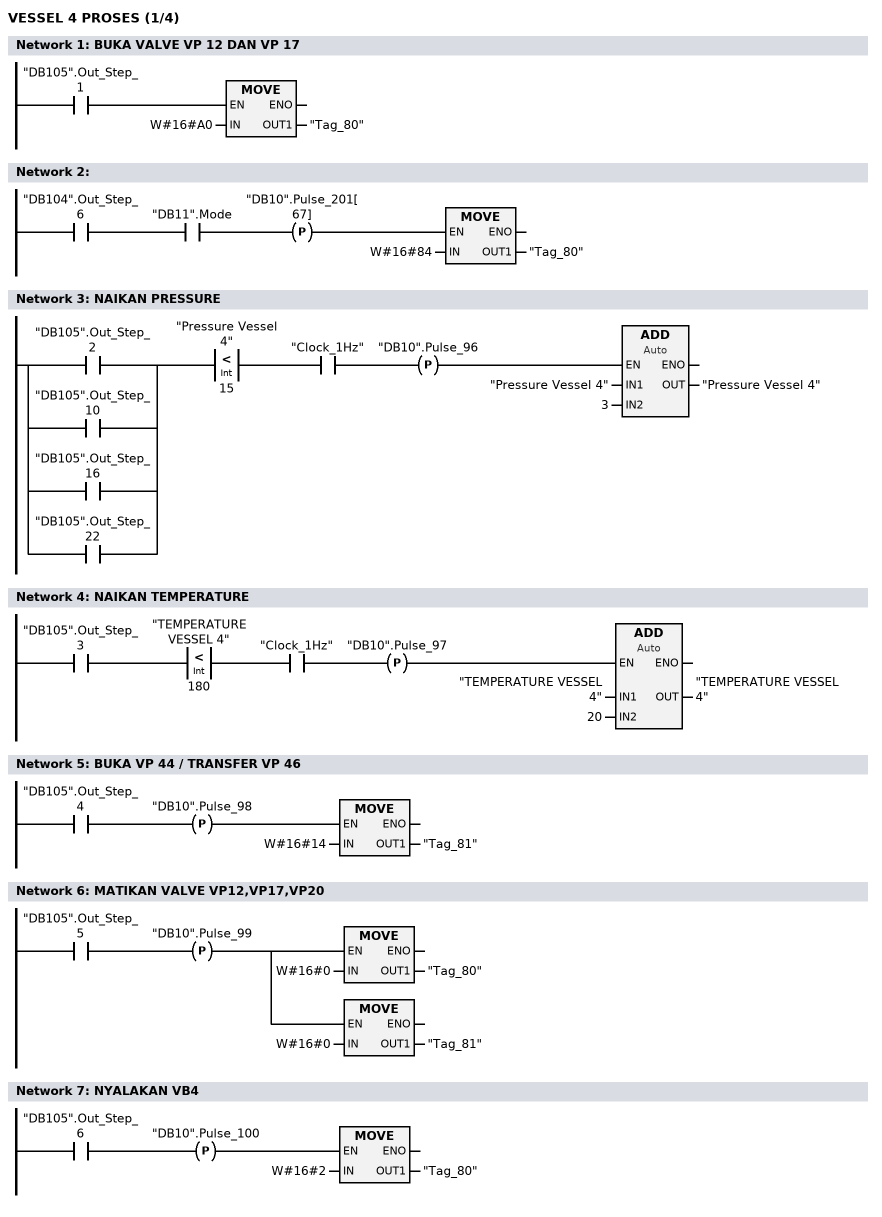
   RUNG wire#powerrail
      Contact( "DB105".Out_Step_1 )
      Move(in := W#16#A0, out1 => "Tag_80")
   END_RUNG
   // the same network as SCL:
   IF "DB105".Out_Step_1 THEN "Tag_80" := W#16#A0; END_IF;
END_REGION

REGION Network 2
   RUNG wire#powerrail
      Contact( "DB104".Out_Step_6 )
      Contact( "DB11".Mode )
      P_Trig( "DB10".Pulse_201[67] )
      Move(in := W#16#84, out1 => "Tag_80")
   END_RUNG
   // the same network as SCL:
   #_w1 := "DB104".Out_Step_6 AND "DB11".Mode;
   #_w2 := #_w1 AND NOT "DB10".Pulse_201[67];   // rising edge
   "DB10".Pulse_201[67] := #_w1;
   IF #_w2 THEN "Tag_80" := W#16#84; END_IF;
END_REGION

REGION Network 3: NAIKAN PRESSURE
   RUNG wire#powerrail
      Contact( "DB105".Out_Step_2 )
      wire#w1
      { S7_Templates := "SrcType := Int" } LT_Contact(in1 := "Pressure Vessel 4", in2 := 15)
      Contact( "Clock_1Hz" )
      P_Trig( "DB10".Pulse_96 )
      Add(in1 := "Pressure Vessel 4", in2 := 3, out => "Pressure Vessel 4")
   END_RUNG
   RUNG wire#powerrail
      Contact( "DB105".Out_Step_10 )
   END_RUNG wire#w1
   RUNG wire#powerrail
      Contact( "DB105".Out_Step_16 )
   END_RUNG wire#w1
   RUNG wire#powerrail
      Contact( "DB105".Out_Step_22 )
   END_RUNG wire#w1
   // the same network as SCL:
   #_w1 := ("DB105".Out_Step_2 OR "DB105".Out_Step_10 OR "DB105".Out_Step_16 OR "DB105".Out_Step_22) AND ("Pressure Vessel 4" < 15) AND "Clock_1Hz";
   #_w2 := #_w1 AND NOT "DB10".Pulse_96;   // rising edge
   "DB10".Pulse_96 := #_w1;
   IF #_w2 THEN "Pressure Vessel 4" := "Pressure Vessel 4" + 3; END_IF;
END_REGION

REGION Network 4: NAIKAN TEMPERATURE
   RUNG wire#powerrail
      Contact( "DB105".Out_Step_3 )
      { S7_Templates := "SrcType := Int" } LT_Contact(in1 := "TEMPERATURE VESSEL 4", in2 := 180)
      Contact( "Clock_1Hz" )
      P_Trig( "DB10".Pulse_97 )
      Add(in1 := "TEMPERATURE VESSEL 4", in2 := 20, out => "TEMPERATURE VESSEL 4")
   END_RUNG
   // the same network as SCL:
   #_w1 := "DB105".Out_Step_3 AND ("TEMPERATURE VESSEL 4" < 180) AND "Clock_1Hz";
   #_w2 := #_w1 AND NOT "DB10".Pulse_97;   // rising edge
   "DB10".Pulse_97 := #_w1;
   IF #_w2 THEN "TEMPERATURE VESSEL 4" := "TEMPERATURE VESSEL 4" + 20; END_IF;
END_REGION

REGION Network 5: BUKA VP 44 / TRANSFER VP 46
   RUNG wire#powerrail
      Contact( "DB105".Out_Step_4 )
      P_Trig( "DB10".Pulse_98 )
      Move(in := W#16#14, out1 => "Tag_81")
   END_RUNG
   // the same network as SCL:
   #_w1 := "DB105".Out_Step_4 AND NOT "DB10".Pulse_98;   // rising edge
   "DB10".Pulse_98 := "DB105".Out_Step_4;
   IF #_w1 THEN "Tag_81" := W#16#14; END_IF;
END_REGION

REGION Network 6: MATIKAN VALVE VP12,VP17,VP20
   RUNG wire#powerrail
      Contact( "DB105".Out_Step_5 )
      P_Trig( "DB10".Pulse_99 )
      wire#w1
      Move(in := W#16#0, out1 => "Tag_80")
   END_RUNG
   RUNG wire#w1
      Move(in := W#16#0, out1 => "Tag_81")
   END_RUNG
   // the same network as SCL:
   #_w1 := "DB105".Out_Step_5 AND NOT "DB10".Pulse_99;   // rising edge
   "DB10".Pulse_99 := "DB105".Out_Step_5;
   IF #_w1 THEN
       "Tag_80" := W#16#0;
       "Tag_81" := W#16#0;
   END_IF;
END_REGION

REGION Network 7: NYALAKAN VB4
   RUNG wire#powerrail
      Contact( "DB105".Out_Step_6 )
      P_Trig( "DB10".Pulse_100 )
      Move(in := W#16#2, out1 => "Tag_80")
   END_RUNG
   // the same network as SCL:
   #_w1 := "DB105".Out_Step_6 AND NOT "DB10".Pulse_100;   // rising edge
   "DB10".Pulse_100 := "DB105".Out_Step_6;
   IF #_w1 THEN "Tag_80" := W#16#2; END_IF;
END_REGION

REGION Network 8: TURUNKAN PRESSURE
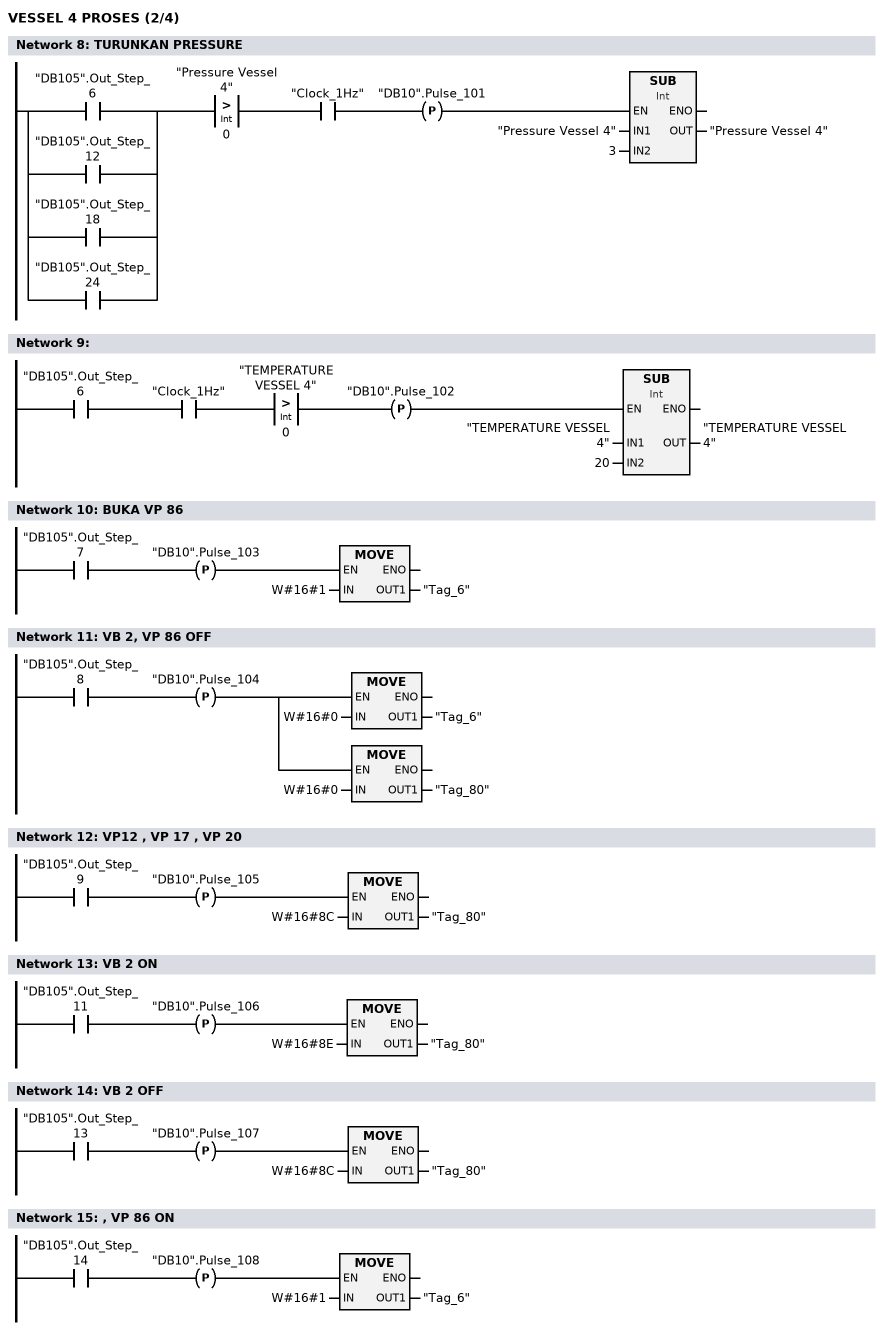
   RUNG wire#powerrail
      Contact( "DB105".Out_Step_6 )
      wire#w1
      { S7_Templates := "SrcType := Int" } GT_Contact(in1 := "Pressure Vessel 4", in2 := 0)
      Contact( "Clock_1Hz" )
      P_Trig( "DB10".Pulse_101 )
      { S7_Templates := "SrcType := Int" } Sub(in1 := "Pressure Vessel 4", in2 := 3, out => "Pressure Vessel 4")
   END_RUNG
   RUNG wire#powerrail
      Contact( "DB105".Out_Step_12 )
   END_RUNG wire#w1
   RUNG wire#powerrail
      Contact( "DB105".Out_Step_18 )
   END_RUNG wire#w1
   RUNG wire#powerrail
      Contact( "DB105".Out_Step_24 )
   END_RUNG wire#w1
   // the same network as SCL:
   #_w1 := ("DB105".Out_Step_6 OR "DB105".Out_Step_12 OR "DB105".Out_Step_18 OR "DB105".Out_Step_24) AND ("Pressure Vessel 4" > 0) AND "Clock_1Hz";
   #_w2 := #_w1 AND NOT "DB10".Pulse_101;   // rising edge
   "DB10".Pulse_101 := #_w1;
   IF #_w2 THEN "Pressure Vessel 4" := "Pressure Vessel 4" - 3; END_IF;
END_REGION

REGION Network 9
   RUNG wire#powerrail
      Contact( "DB105".Out_Step_6 )
      Contact( "Clock_1Hz" )
      { S7_Templates := "SrcType := Int" } GT_Contact(in1 := "TEMPERATURE VESSEL 4", in2 := 0)
      P_Trig( "DB10".Pulse_102 )
      { S7_Templates := "SrcType := Int" } Sub(in1 := "TEMPERATURE VESSEL 4", in2 := 20, out => "TEMPERATURE VESSEL 4")
   END_RUNG
   // the same network as SCL:
   #_w1 := "DB105".Out_Step_6 AND "Clock_1Hz" AND ("TEMPERATURE VESSEL 4" > 0);
   #_w2 := #_w1 AND NOT "DB10".Pulse_102;   // rising edge
   "DB10".Pulse_102 := #_w1;
   IF #_w2 THEN "TEMPERATURE VESSEL 4" := "TEMPERATURE VESSEL 4" - 20; END_IF;
END_REGION

REGION Network 10: BUKA VP 86
   RUNG wire#powerrail
      Contact( "DB105".Out_Step_7 )
      P_Trig( "DB10".Pulse_103 )
      Move(in := W#16#1, out1 => "Tag_6")
   END_RUNG
   // the same network as SCL:
   #_w1 := "DB105".Out_Step_7 AND NOT "DB10".Pulse_103;   // rising edge
   "DB10".Pulse_103 := "DB105".Out_Step_7;
   IF #_w1 THEN "Tag_6" := W#16#1; END_IF;
END_REGION

REGION Network 11: VB 2, VP 86 OFF
   RUNG wire#powerrail
      Contact( "DB105".Out_Step_8 )
      P_Trig( "DB10".Pulse_104 )
      wire#w1
      Move(in := W#16#0, out1 => "Tag_6")
   END_RUNG
   RUNG wire#w1
      Move(in := W#16#0, out1 => "Tag_80")
   END_RUNG
   // the same network as SCL:
   #_w1 := "DB105".Out_Step_8 AND NOT "DB10".Pulse_104;   // rising edge
   "DB10".Pulse_104 := "DB105".Out_Step_8;
   IF #_w1 THEN
       "Tag_6" := W#16#0;
       "Tag_80" := W#16#0;
   END_IF;
END_REGION

REGION Network 12: VP12 , VP 17 , VP 20
   RUNG wire#powerrail
      Contact( "DB105".Out_Step_9 )
      P_Trig( "DB10".Pulse_105 )
      Move(in := W#16#8C, out1 => "Tag_80")
   END_RUNG
   // the same network as SCL:
   #_w1 := "DB105".Out_Step_9 AND NOT "DB10".Pulse_105;   // rising edge
   "DB10".Pulse_105 := "DB105".Out_Step_9;
   IF #_w1 THEN "Tag_80" := W#16#8C; END_IF;
END_REGION

REGION Network 13: VB 2 ON
   RUNG wire#powerrail
      Contact( "DB105".Out_Step_11 )
      P_Trig( "DB10".Pulse_106 )
      Move(in := W#16#8E, out1 => "Tag_80")
   END_RUNG
   // the same network as SCL:
   #_w1 := "DB105".Out_Step_11 AND NOT "DB10".Pulse_106;   // rising edge
   "DB10".Pulse_106 := "DB105".Out_Step_11;
   IF #_w1 THEN "Tag_80" := W#16#8E; END_IF;
END_REGION

REGION Network 14: VB 2 OFF
   RUNG wire#powerrail
      Contact( "DB105".Out_Step_13 )
      P_Trig( "DB10".Pulse_107 )
      Move(in := W#16#8C, out1 => "Tag_80")
   END_RUNG
   // the same network as SCL:
   #_w1 := "DB105".Out_Step_13 AND NOT "DB10".Pulse_107;   // rising edge
   "DB10".Pulse_107 := "DB105".Out_Step_13;
   IF #_w1 THEN "Tag_80" := W#16#8C; END_IF;
END_REGION

REGION Network 15: , VP 86 ON
   RUNG wire#powerrail
      Contact( "DB105".Out_Step_14 )
      P_Trig( "DB10".Pulse_108 )
      Move(in := W#16#1, out1 => "Tag_6")
   END_RUNG
   // the same network as SCL:
   #_w1 := "DB105".Out_Step_14 AND NOT "DB10".Pulse_108;   // rising edge
   "DB10".Pulse_108 := "DB105".Out_Step_14;
   IF #_w1 THEN "Tag_6" := W#16#1; END_IF;
END_REGION

REGION Network 16: VP 86 OFF
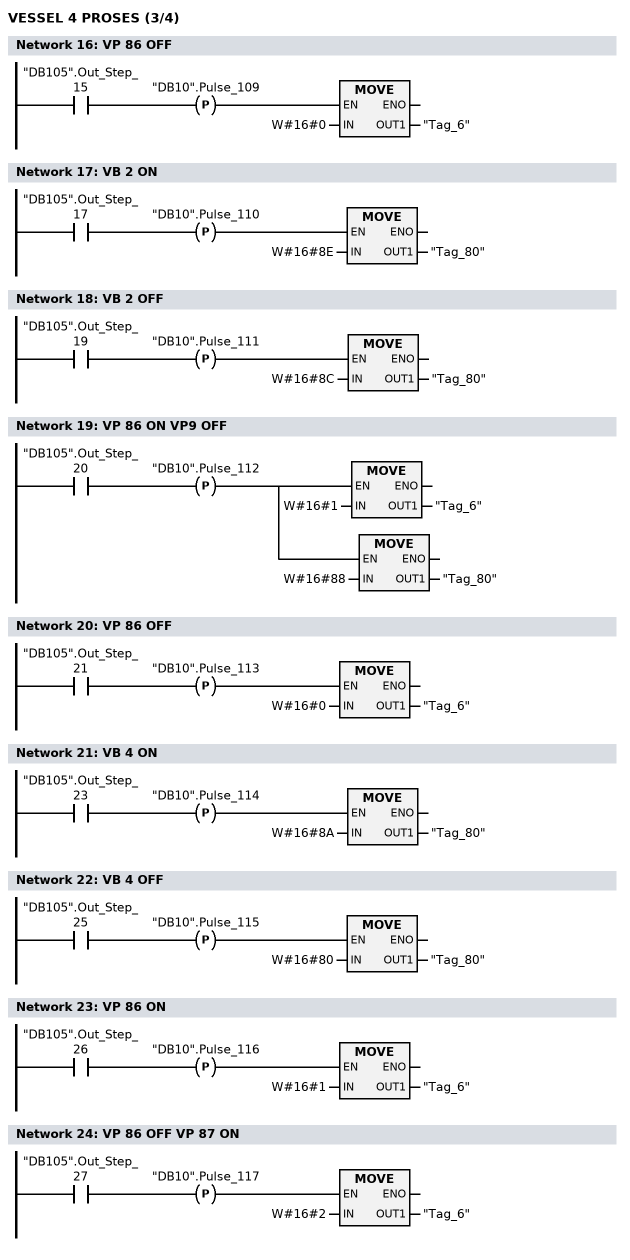
   RUNG wire#powerrail
      Contact( "DB105".Out_Step_15 )
      P_Trig( "DB10".Pulse_109 )
      Move(in := W#16#0, out1 => "Tag_6")
   END_RUNG
   // the same network as SCL:
   #_w1 := "DB105".Out_Step_15 AND NOT "DB10".Pulse_109;   // rising edge
   "DB10".Pulse_109 := "DB105".Out_Step_15;
   IF #_w1 THEN "Tag_6" := W#16#0; END_IF;
END_REGION

REGION Network 17: VB 2 ON
   RUNG wire#powerrail
      Contact( "DB105".Out_Step_17 )
      P_Trig( "DB10".Pulse_110 )
      Move(in := W#16#8E, out1 => "Tag_80")
   END_RUNG
   // the same network as SCL:
   #_w1 := "DB105".Out_Step_17 AND NOT "DB10".Pulse_110;   // rising edge
   "DB10".Pulse_110 := "DB105".Out_Step_17;
   IF #_w1 THEN "Tag_80" := W#16#8E; END_IF;
END_REGION

REGION Network 18: VB 2 OFF
   RUNG wire#powerrail
      Contact( "DB105".Out_Step_19 )
      P_Trig( "DB10".Pulse_111 )
      Move(in := W#16#8C, out1 => "Tag_80")
   END_RUNG
   // the same network as SCL:
   #_w1 := "DB105".Out_Step_19 AND NOT "DB10".Pulse_111;   // rising edge
   "DB10".Pulse_111 := "DB105".Out_Step_19;
   IF #_w1 THEN "Tag_80" := W#16#8C; END_IF;
END_REGION

REGION Network 19: VP 86 ON VP9 OFF
   RUNG wire#powerrail
      Contact( "DB105".Out_Step_20 )
      P_Trig( "DB10".Pulse_112 )
      wire#w1
      Move(in := W#16#1, out1 => "Tag_6")
   END_RUNG
   RUNG wire#w1
      Move(in := W#16#88, out1 => "Tag_80")
   END_RUNG
   // the same network as SCL:
   #_w1 := "DB105".Out_Step_20 AND NOT "DB10".Pulse_112;   // rising edge
   "DB10".Pulse_112 := "DB105".Out_Step_20;
   IF #_w1 THEN
       "Tag_6" := W#16#1;
       "Tag_80" := W#16#88;
   END_IF;
END_REGION

REGION Network 20: VP 86 OFF
   RUNG wire#powerrail
      Contact( "DB105".Out_Step_21 )
      P_Trig( "DB10".Pulse_113 )
      Move(in := W#16#0, out1 => "Tag_6")
   END_RUNG
   // the same network as SCL:
   #_w1 := "DB105".Out_Step_21 AND NOT "DB10".Pulse_113;   // rising edge
   "DB10".Pulse_113 := "DB105".Out_Step_21;
   IF #_w1 THEN "Tag_6" := W#16#0; END_IF;
END_REGION

REGION Network 21: VB 4 ON
   RUNG wire#powerrail
      Contact( "DB105".Out_Step_23 )
      P_Trig( "DB10".Pulse_114 )
      Move(in := W#16#8A, out1 => "Tag_80")
   END_RUNG
   // the same network as SCL:
   #_w1 := "DB105".Out_Step_23 AND NOT "DB10".Pulse_114;   // rising edge
   "DB10".Pulse_114 := "DB105".Out_Step_23;
   IF #_w1 THEN "Tag_80" := W#16#8A; END_IF;
END_REGION

REGION Network 22: VB 4 OFF
   RUNG wire#powerrail
      Contact( "DB105".Out_Step_25 )
      P_Trig( "DB10".Pulse_115 )
      Move(in := W#16#80, out1 => "Tag_80")
   END_RUNG
   // the same network as SCL:
   #_w1 := "DB105".Out_Step_25 AND NOT "DB10".Pulse_115;   // rising edge
   "DB10".Pulse_115 := "DB105".Out_Step_25;
   IF #_w1 THEN "Tag_80" := W#16#80; END_IF;
END_REGION

REGION Network 23: VP 86 ON
   RUNG wire#powerrail
      Contact( "DB105".Out_Step_26 )
      P_Trig( "DB10".Pulse_116 )
      Move(in := W#16#1, out1 => "Tag_6")
   END_RUNG
   // the same network as SCL:
   #_w1 := "DB105".Out_Step_26 AND NOT "DB10".Pulse_116;   // rising edge
   "DB10".Pulse_116 := "DB105".Out_Step_26;
   IF #_w1 THEN "Tag_6" := W#16#1; END_IF;
END_REGION

REGION Network 24: VP 86 OFF VP 87 ON
   RUNG wire#powerrail
      Contact( "DB105".Out_Step_27 )
      P_Trig( "DB10".Pulse_117 )
      Move(in := W#16#2, out1 => "Tag_6")
   END_RUNG
   // the same network as SCL:
   #_w1 := "DB105".Out_Step_27 AND NOT "DB10".Pulse_117;   // rising edge
   "DB10".Pulse_117 := "DB105".Out_Step_27;
   IF #_w1 THEN "Tag_6" := W#16#2; END_IF;
END_REGION

REGION Network 25: VP 87 OFF
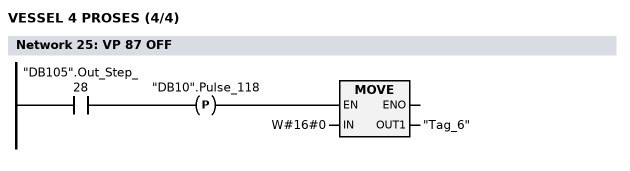
   RUNG wire#powerrail
      Contact( "DB105".Out_Step_28 )
      P_Trig( "DB10".Pulse_118 )
      Move(in := W#16#0, out1 => "Tag_6")
   END_RUNG
   // the same network as SCL:
   #_w1 := "DB105".Out_Step_28 AND NOT "DB10".Pulse_118;   // rising edge
   "DB10".Pulse_118 := "DB105".Out_Step_28;
   IF #_w1 THEN "Tag_6" := W#16#0; END_IF;
END_REGION
END_FUNCTION

FUNCTION "SEQUENCE V4 PROSES" : Void   // FC16, LAD
{ S7_Optimized_Access := 'TRUE' }
VERSION : 0.1
   VAR_TEMP   // added for the SCL form of the ladder/FBD networks
      _w1 : Bool;
      _w2 : Bool;
      _s5time1 : S5Time;
   END_VAR
BEGIN

REGION Network 1: START PROSES
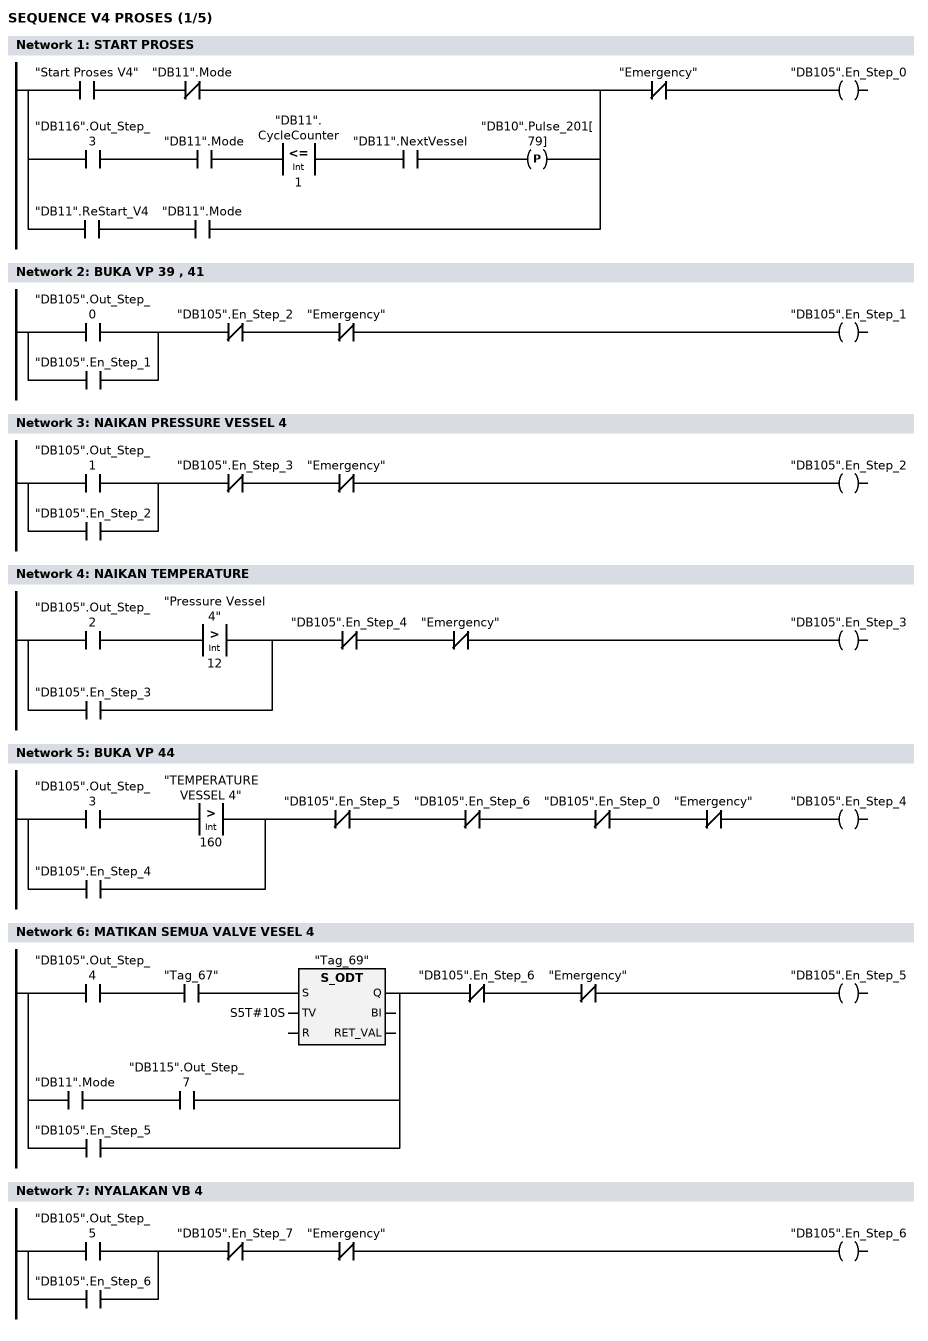
   RUNG wire#powerrail
      Contact( "Start Proses V4" )
      I_Contact( "DB11".Mode )
      wire#w1
      I_Contact( "Emergency" )
      Coil( "DB105".En_Step_0 )
   END_RUNG
   RUNG wire#powerrail
      Contact( "DB116".Out_Step_3 )
      Contact( "DB11".Mode )
      { S7_Templates := "SrcType := Int" } LE_Contact(in1 := "DB11".CycleCounter, in2 := 1)
      Contact( "DB11".NextVessel )
      P_Trig( "DB10".Pulse_201[79] )
   END_RUNG wire#w1
   RUNG wire#powerrail
      Contact( "DB11".ReStart_V4 )
      Contact( "DB11".Mode )
   END_RUNG wire#w1
   // the same network as SCL:
   #_w1 := "DB116".Out_Step_3 AND "DB11".Mode AND ("DB11".CycleCounter <= 1) AND "DB11".NextVessel;
   #_w2 := #_w1 AND NOT "DB10".Pulse_201[79];   // rising edge
   "DB10".Pulse_201[79] := #_w1;
   "DB105".En_Step_0 := (("Start Proses V4" AND NOT "DB11".Mode) OR #_w2 OR ("DB11".ReStart_V4 AND "DB11".Mode)) AND NOT "Emergency";
END_REGION

REGION Network 2: BUKA VP 39 , 41
   RUNG wire#powerrail
      Contact( "DB105".Out_Step_0 )
      wire#w1
      I_Contact( "DB105".En_Step_2 )
      I_Contact( "Emergency" )
      Coil( "DB105".En_Step_1 )
   END_RUNG
   RUNG wire#powerrail
      Contact( "DB105".En_Step_1 )
   END_RUNG wire#w1
   // the same network as SCL:
   "DB105".En_Step_1 := ("DB105".Out_Step_0 OR "DB105".En_Step_1) AND NOT "DB105".En_Step_2 AND NOT "Emergency";
END_REGION

REGION Network 3: NAIKAN PRESSURE VESSEL 4
   RUNG wire#powerrail
      Contact( "DB105".Out_Step_1 )
      wire#w1
      I_Contact( "DB105".En_Step_3 )
      I_Contact( "Emergency" )
      Coil( "DB105".En_Step_2 )
   END_RUNG
   RUNG wire#powerrail
      Contact( "DB105".En_Step_2 )
   END_RUNG wire#w1
   // the same network as SCL:
   "DB105".En_Step_2 := ("DB105".Out_Step_1 OR "DB105".En_Step_2) AND NOT "DB105".En_Step_3 AND NOT "Emergency";
END_REGION

REGION Network 4: NAIKAN TEMPERATURE
   RUNG wire#powerrail
      Contact( "DB105".Out_Step_2 )
      { S7_Templates := "SrcType := Int" } GT_Contact(in1 := "Pressure Vessel 4", in2 := 12)
      wire#w1
      I_Contact( "DB105".En_Step_4 )
      I_Contact( "Emergency" )
      Coil( "DB105".En_Step_3 )
   END_RUNG
   RUNG wire#powerrail
      Contact( "DB105".En_Step_3 )
   END_RUNG wire#w1
   // the same network as SCL:
   "DB105".En_Step_3 := (("DB105".Out_Step_2 AND ("Pressure Vessel 4" > 12)) OR "DB105".En_Step_3) AND NOT "DB105".En_Step_4 AND NOT "Emergency";
END_REGION

REGION Network 5: BUKA VP 44
   RUNG wire#powerrail
      Contact( "DB105".Out_Step_3 )
      { S7_Templates := "SrcType := Int" } GT_Contact(in1 := "TEMPERATURE VESSEL 4", in2 := 160)
      wire#w1
      I_Contact( "DB105".En_Step_5 )
      I_Contact( "DB105".En_Step_6 )
      I_Contact( "DB105".En_Step_0 )
      I_Contact( "Emergency" )
      Coil( "DB105".En_Step_4 )
   END_RUNG
   RUNG wire#powerrail
      Contact( "DB105".En_Step_4 )
   END_RUNG wire#w1
   // the same network as SCL:
   "DB105".En_Step_4 := (("DB105".Out_Step_3 AND ("TEMPERATURE VESSEL 4" > 160)) OR "DB105".En_Step_4) AND NOT "DB105".En_Step_5 AND NOT "DB105".En_Step_6 AND NOT "DB105".En_Step_0 AND NOT "Emergency";
END_REGION

REGION Network 6: MATIKAN SEMUA VALVE VESEL 4
   RUNG wire#powerrail
      Contact( "DB105".Out_Step_4 )
      Contact( "Tag_67" )
      S_ODT(T_NO := "Tag_69", TV := S5T#10S, R :=, BI =>, RET_VAL =>)
      wire#w1
      I_Contact( "DB105".En_Step_6 )
      I_Contact( "Emergency" )
      Coil( "DB105".En_Step_5 )
   END_RUNG
   RUNG wire#powerrail
      Contact( "DB11".Mode )
      Contact( "DB115".Out_Step_7 )
   END_RUNG wire#w1
   RUNG wire#powerrail
      Contact( "DB105".En_Step_5 )
   END_RUNG wire#w1
   // the same network as SCL:
   #_s5time1 := S_ODT(T_NO := "Tag_69", S := "DB105".Out_Step_4 AND "Tag_67", TV := S5T#10S, Q => #_w1);
   "DB105".En_Step_5 := (#_w1 OR ("DB11".Mode AND "DB115".Out_Step_7) OR "DB105".En_Step_5) AND NOT "DB105".En_Step_6 AND NOT "Emergency";
END_REGION

REGION Network 7: NYALAKAN VB 4
   RUNG wire#powerrail
      Contact( "DB105".Out_Step_5 )
      wire#w1
      I_Contact( "DB105".En_Step_7 )
      I_Contact( "Emergency" )
      Coil( "DB105".En_Step_6 )
   END_RUNG
   RUNG wire#powerrail
      Contact( "DB105".En_Step_6 )
   END_RUNG wire#w1
   // the same network as SCL:
   "DB105".En_Step_6 := ("DB105".Out_Step_5 OR "DB105".En_Step_6) AND NOT "DB105".En_Step_7 AND NOT "Emergency";
END_REGION

REGION Network 8
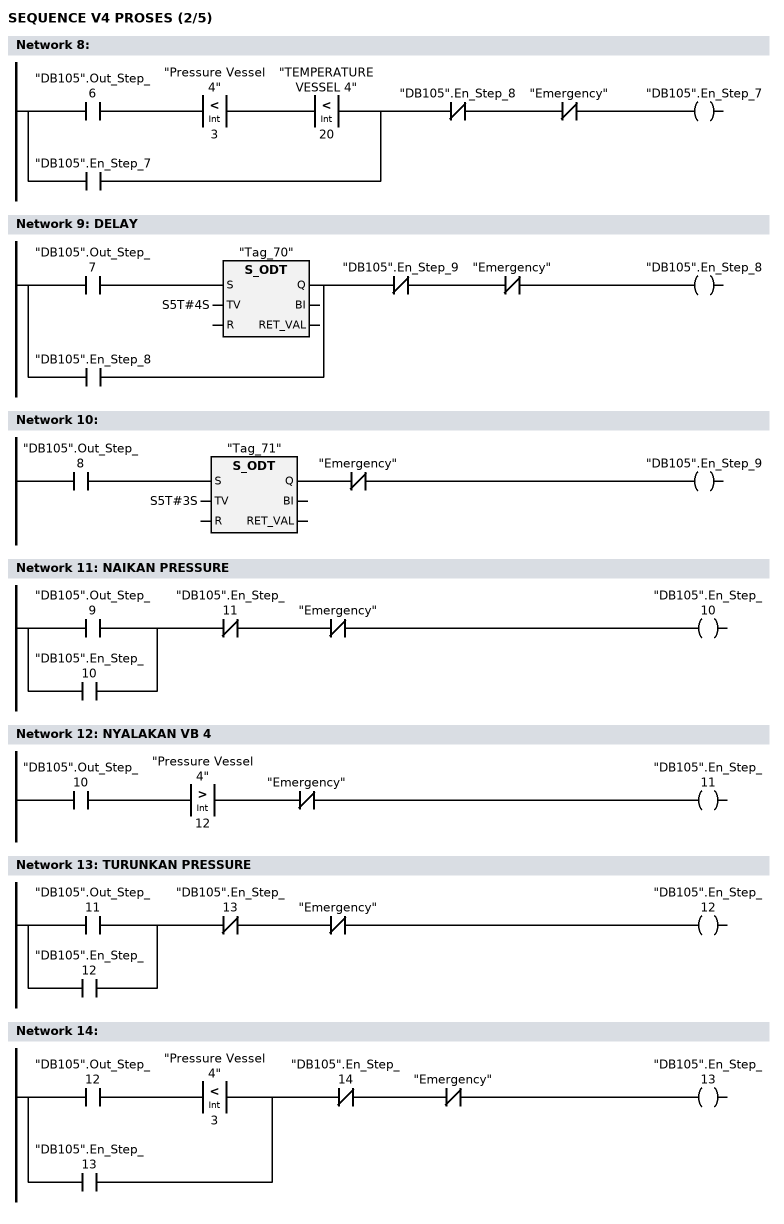
   RUNG wire#powerrail
      Contact( "DB105".Out_Step_6 )
      { S7_Templates := "SrcType := Int" } LT_Contact(in1 := "Pressure Vessel 4", in2 := 3)
      { S7_Templates := "SrcType := Int" } LT_Contact(in1 := "TEMPERATURE VESSEL 4", in2 := 20)
      wire#w1
      I_Contact( "DB105".En_Step_8 )
      I_Contact( "Emergency" )
      Coil( "DB105".En_Step_7 )
   END_RUNG
   RUNG wire#powerrail
      Contact( "DB105".En_Step_7 )
   END_RUNG wire#w1
   // the same network as SCL:
   "DB105".En_Step_7 := (("DB105".Out_Step_6 AND ("Pressure Vessel 4" < 3) AND ("TEMPERATURE VESSEL 4" < 20)) OR "DB105".En_Step_7) AND NOT "DB105".En_Step_8 AND NOT "Emergency";
END_REGION

REGION Network 9: DELAY
   RUNG wire#powerrail
      Contact( "DB105".Out_Step_7 )
      S_ODT(T_NO := "Tag_70", TV := S5T#4S, R :=, BI =>, RET_VAL =>)
      wire#w1
      I_Contact( "DB105".En_Step_9 )
      I_Contact( "Emergency" )
      Coil( "DB105".En_Step_8 )
   END_RUNG
   RUNG wire#powerrail
      Contact( "DB105".En_Step_8 )
   END_RUNG wire#w1
   // the same network as SCL:
   #_s5time1 := S_ODT(T_NO := "Tag_70", S := "DB105".Out_Step_7, TV := S5T#4S, Q => #_w1);
   "DB105".En_Step_8 := (#_w1 OR "DB105".En_Step_8) AND NOT "DB105".En_Step_9 AND NOT "Emergency";
END_REGION

REGION Network 10
   RUNG wire#powerrail
      Contact( "DB105".Out_Step_8 )
      S_ODT(T_NO := "Tag_71", TV := S5T#3S, R :=, BI =>, RET_VAL =>)
      I_Contact( "Emergency" )
      Coil( "DB105".En_Step_9 )
   END_RUNG
   // the same network as SCL:
   #_s5time1 := S_ODT(T_NO := "Tag_71", S := "DB105".Out_Step_8, TV := S5T#3S, Q => #_w1);
   "DB105".En_Step_9 := #_w1 AND NOT "Emergency";
END_REGION

REGION Network 11: NAIKAN PRESSURE
   RUNG wire#powerrail
      Contact( "DB105".Out_Step_9 )
      wire#w1
      I_Contact( "DB105".En_Step_11 )
      I_Contact( "Emergency" )
      Coil( "DB105".En_Step_10 )
   END_RUNG
   RUNG wire#powerrail
      Contact( "DB105".En_Step_10 )
   END_RUNG wire#w1
   // the same network as SCL:
   "DB105".En_Step_10 := ("DB105".Out_Step_9 OR "DB105".En_Step_10) AND NOT "DB105".En_Step_11 AND NOT "Emergency";
END_REGION

REGION Network 12: NYALAKAN VB 4
   RUNG wire#powerrail
      Contact( "DB105".Out_Step_10 )
      { S7_Templates := "SrcType := Int" } GT_Contact(in1 := "Pressure Vessel 4", in2 := 12)
      I_Contact( "Emergency" )
      Coil( "DB105".En_Step_11 )
   END_RUNG
   // the same network as SCL:
   "DB105".En_Step_11 := "DB105".Out_Step_10 AND ("Pressure Vessel 4" > 12) AND NOT "Emergency";
END_REGION

REGION Network 13: TURUNKAN PRESSURE
   RUNG wire#powerrail
      Contact( "DB105".Out_Step_11 )
      wire#w1
      I_Contact( "DB105".En_Step_13 )
      I_Contact( "Emergency" )
      Coil( "DB105".En_Step_12 )
   END_RUNG
   RUNG wire#powerrail
      Contact( "DB105".En_Step_12 )
   END_RUNG wire#w1
   // the same network as SCL:
   "DB105".En_Step_12 := ("DB105".Out_Step_11 OR "DB105".En_Step_12) AND NOT "DB105".En_Step_13 AND NOT "Emergency";
END_REGION

REGION Network 14
   RUNG wire#powerrail
      Contact( "DB105".Out_Step_12 )
      { S7_Templates := "SrcType := Int" } LT_Contact(in1 := "Pressure Vessel 4", in2 := 3)
      wire#w1
      I_Contact( "DB105".En_Step_14 )
      I_Contact( "Emergency" )
      Coil( "DB105".En_Step_13 )
   END_RUNG
   RUNG wire#powerrail
      Contact( "DB105".En_Step_13 )
   END_RUNG wire#w1
   // the same network as SCL:
   "DB105".En_Step_13 := (("DB105".Out_Step_12 AND ("Pressure Vessel 4" < 3)) OR "DB105".En_Step_13) AND NOT "DB105".En_Step_14 AND NOT "Emergency";
END_REGION

REGION Network 15
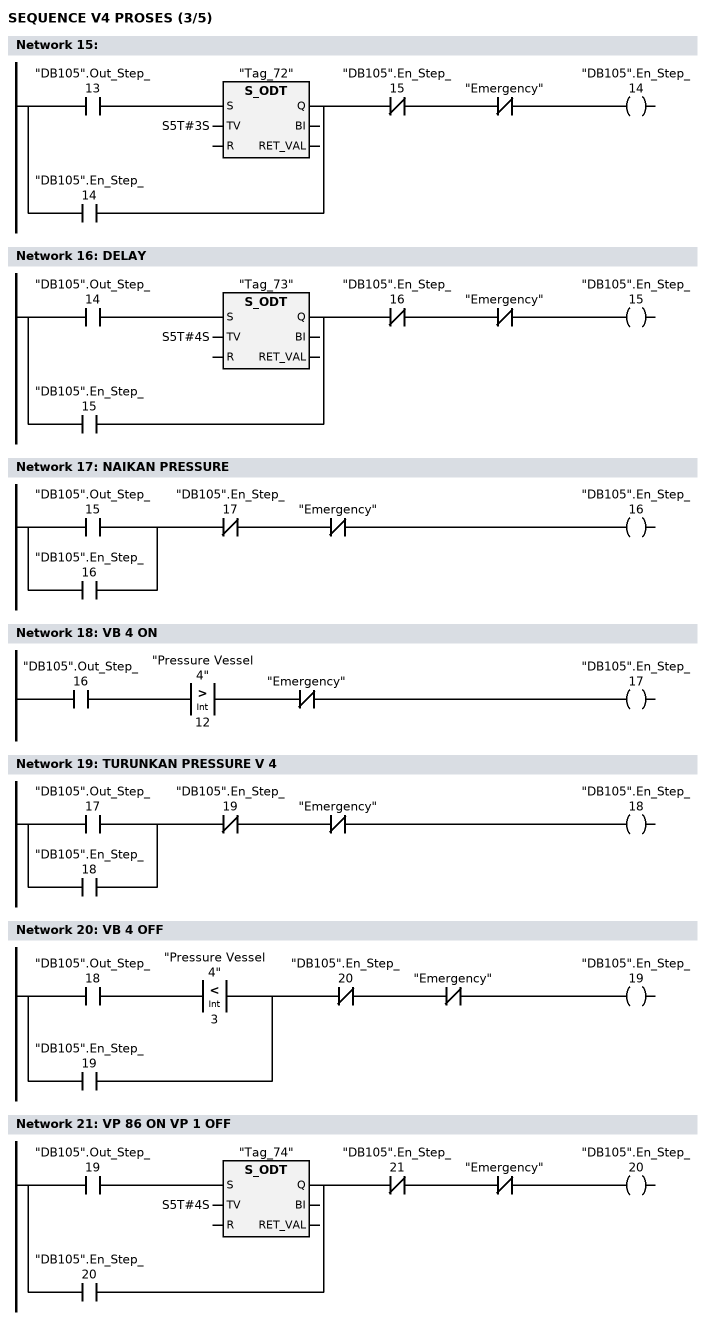
   RUNG wire#powerrail
      Contact( "DB105".Out_Step_13 )
      S_ODT(T_NO := "Tag_72", TV := S5T#3S, R :=, BI =>, RET_VAL =>)
      wire#w1
      I_Contact( "DB105".En_Step_15 )
      I_Contact( "Emergency" )
      Coil( "DB105".En_Step_14 )
   END_RUNG
   RUNG wire#powerrail
      Contact( "DB105".En_Step_14 )
   END_RUNG wire#w1
   // the same network as SCL:
   #_s5time1 := S_ODT(T_NO := "Tag_72", S := "DB105".Out_Step_13, TV := S5T#3S, Q => #_w1);
   "DB105".En_Step_14 := (#_w1 OR "DB105".En_Step_14) AND NOT "DB105".En_Step_15 AND NOT "Emergency";
END_REGION

REGION Network 16: DELAY
   RUNG wire#powerrail
      Contact( "DB105".Out_Step_14 )
      S_ODT(T_NO := "Tag_73", TV := S5T#4S, R :=, BI =>, RET_VAL =>)
      wire#w1
      I_Contact( "DB105".En_Step_16 )
      I_Contact( "Emergency" )
      Coil( "DB105".En_Step_15 )
   END_RUNG
   RUNG wire#powerrail
      Contact( "DB105".En_Step_15 )
   END_RUNG wire#w1
   // the same network as SCL:
   #_s5time1 := S_ODT(T_NO := "Tag_73", S := "DB105".Out_Step_14, TV := S5T#4S, Q => #_w1);
   "DB105".En_Step_15 := (#_w1 OR "DB105".En_Step_15) AND NOT "DB105".En_Step_16 AND NOT "Emergency";
END_REGION

REGION Network 17: NAIKAN PRESSURE
   RUNG wire#powerrail
      Contact( "DB105".Out_Step_15 )
      wire#w1
      I_Contact( "DB105".En_Step_17 )
      I_Contact( "Emergency" )
      Coil( "DB105".En_Step_16 )
   END_RUNG
   RUNG wire#powerrail
      Contact( "DB105".En_Step_16 )
   END_RUNG wire#w1
   // the same network as SCL:
   "DB105".En_Step_16 := ("DB105".Out_Step_15 OR "DB105".En_Step_16) AND NOT "DB105".En_Step_17 AND NOT "Emergency";
END_REGION

REGION Network 18: VB 4 ON
   RUNG wire#powerrail
      Contact( "DB105".Out_Step_16 )
      { S7_Templates := "SrcType := Int" } GT_Contact(in1 := "Pressure Vessel 4", in2 := 12)
      I_Contact( "Emergency" )
      Coil( "DB105".En_Step_17 )
   END_RUNG
   // the same network as SCL:
   "DB105".En_Step_17 := "DB105".Out_Step_16 AND ("Pressure Vessel 4" > 12) AND NOT "Emergency";
END_REGION

REGION Network 19: TURUNKAN PRESSURE V 4
   RUNG wire#powerrail
      Contact( "DB105".Out_Step_17 )
      wire#w1
      I_Contact( "DB105".En_Step_19 )
      I_Contact( "Emergency" )
      Coil( "DB105".En_Step_18 )
   END_RUNG
   RUNG wire#powerrail
      Contact( "DB105".En_Step_18 )
   END_RUNG wire#w1
   // the same network as SCL:
   "DB105".En_Step_18 := ("DB105".Out_Step_17 OR "DB105".En_Step_18) AND NOT "DB105".En_Step_19 AND NOT "Emergency";
END_REGION

REGION Network 20: VB 4 OFF
   RUNG wire#powerrail
      Contact( "DB105".Out_Step_18 )
      { S7_Templates := "SrcType := Int" } LT_Contact(in1 := "Pressure Vessel 4", in2 := 3)
      wire#w1
      I_Contact( "DB105".En_Step_20 )
      I_Contact( "Emergency" )
      Coil( "DB105".En_Step_19 )
   END_RUNG
   RUNG wire#powerrail
      Contact( "DB105".En_Step_19 )
   END_RUNG wire#w1
   // the same network as SCL:
   "DB105".En_Step_19 := (("DB105".Out_Step_18 AND ("Pressure Vessel 4" < 3)) OR "DB105".En_Step_19) AND NOT "DB105".En_Step_20 AND NOT "Emergency";
END_REGION

REGION Network 21: VP 86 ON VP 1 OFF
   RUNG wire#powerrail
      Contact( "DB105".Out_Step_19 )
      S_ODT(T_NO := "Tag_74", TV := S5T#4S, R :=, BI =>, RET_VAL =>)
      wire#w1
      I_Contact( "DB105".En_Step_21 )
      I_Contact( "Emergency" )
      Coil( "DB105".En_Step_20 )
   END_RUNG
   RUNG wire#powerrail
      Contact( "DB105".En_Step_20 )
   END_RUNG wire#w1
   // the same network as SCL:
   #_s5time1 := S_ODT(T_NO := "Tag_74", S := "DB105".Out_Step_19, TV := S5T#4S, Q => #_w1);
   "DB105".En_Step_20 := (#_w1 OR "DB105".En_Step_20) AND NOT "DB105".En_Step_21 AND NOT "Emergency";
END_REGION

REGION Network 22: VP 86 OFF VP 87 ON
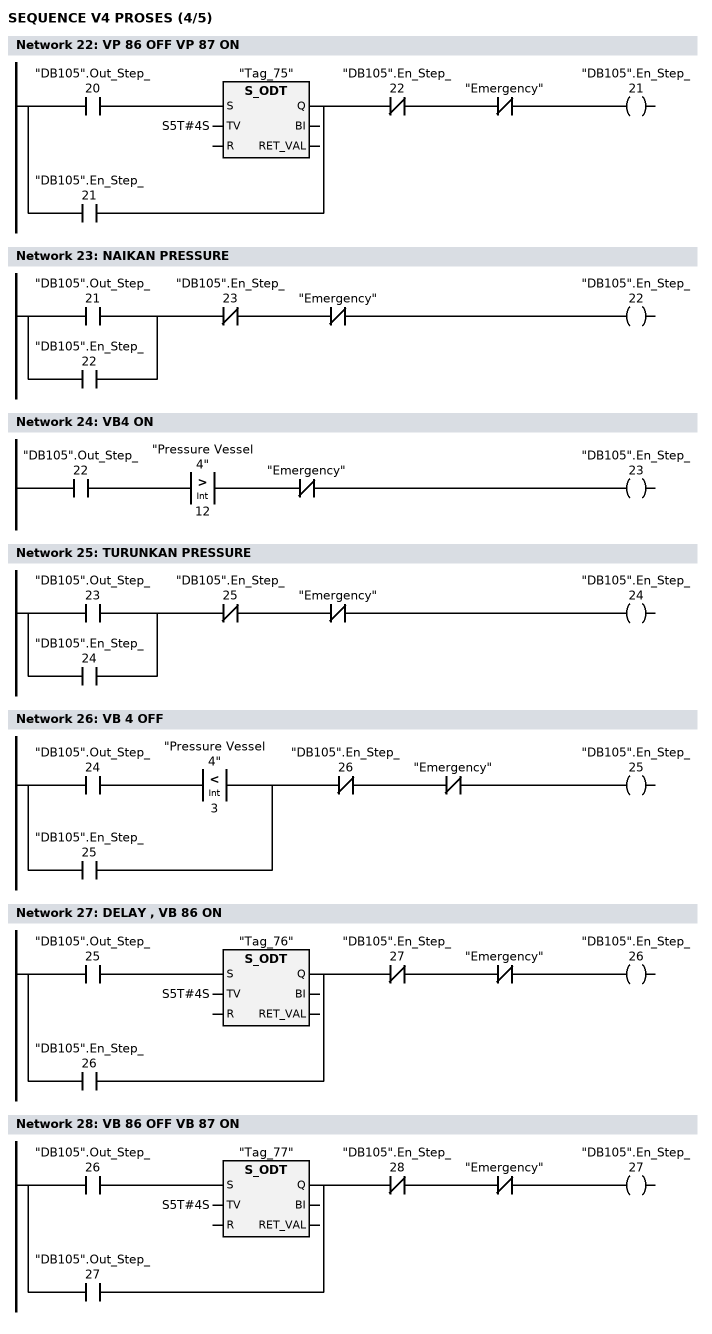
   RUNG wire#powerrail
      Contact( "DB105".Out_Step_20 )
      S_ODT(T_NO := "Tag_75", TV := S5T#4S, R :=, BI =>, RET_VAL =>)
      wire#w1
      I_Contact( "DB105".En_Step_22 )
      I_Contact( "Emergency" )
      Coil( "DB105".En_Step_21 )
   END_RUNG
   RUNG wire#powerrail
      Contact( "DB105".En_Step_21 )
   END_RUNG wire#w1
   // the same network as SCL:
   #_s5time1 := S_ODT(T_NO := "Tag_75", S := "DB105".Out_Step_20, TV := S5T#4S, Q => #_w1);
   "DB105".En_Step_21 := (#_w1 OR "DB105".En_Step_21) AND NOT "DB105".En_Step_22 AND NOT "Emergency";
END_REGION
